// TIA Portal project "SSA-3GHz_V18" (V18) (continued)
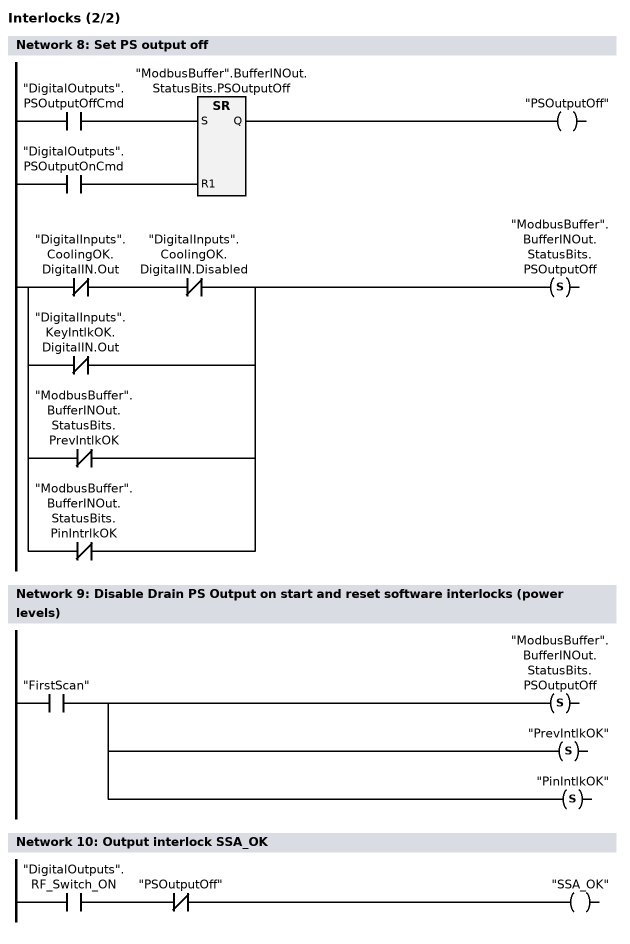
   RUNG wire#powerrail
      Contact( "DigitalOutputs".PSOutputOffCmd )
      S_SR(operand := "ModbusBuffer".BufferINOut.StatusBits.PSOutputOff, r1 := wire#w1)
      Coil( "PSOutputOff" )
   END_RUNG
   RUNG wire#powerrail
      Contact( "DigitalOutputs".PSOutputOnCmd )
   END_RUNG wire#w1
   RUNG wire#powerrail
      I_Contact( "DigitalInputs".CoolingOK.DigitalIN.Out )
      I_Contact( "DigitalInputs".CoolingOK.DigitalIN.Disabled )
      wire#w2
      S_Coil( "ModbusBuffer".BufferINOut.StatusBits.PSOutputOff )
   END_RUNG
   RUNG wire#powerrail
      I_Contact( "DigitalInputs".KeyIntlkOK.DigitalIN.Out )
   END_RUNG wire#w2
   RUNG wire#powerrail
      I_Contact( "ModbusBuffer".BufferINOut.StatusBits.PrevIntlkOK )
   END_RUNG wire#w2
   RUNG wire#powerrail
      I_Contact( "ModbusBuffer".BufferINOut.StatusBits.PinIntrlkOK )
   END_RUNG wire#w2
   // the same network as SCL:
   IF "DigitalOutputs".PSOutputOffCmd THEN
       "ModbusBuffer".BufferINOut.StatusBits.PSOutputOff := TRUE;   // SR flip-flop
   END_IF;
   IF "DigitalOutputs".PSOutputOnCmd THEN "ModbusBuffer".BufferINOut.StatusBits.PSOutputOff := FALSE; END_IF;
   "PSOutputOff" := "ModbusBuffer".BufferINOut.StatusBits.PSOutputOff;
   IF (NOT "DigitalInputs".CoolingOK.DigitalIN.Out AND NOT "DigitalInputs".CoolingOK.DigitalIN.Disabled) OR NOT "DigitalInputs".KeyIntlkOK.DigitalIN.Out OR NOT "ModbusBuffer".BufferINOut.StatusBits.PrevIntlkOK OR NOT "ModbusBuffer".BufferINOut.StatusBits.PinIntrlkOK THEN
       "ModbusBuffer".BufferINOut.StatusBits.PSOutputOff := TRUE;
   END_IF;
END_REGION

REGION Network 9: Disable Drain PS Output on start and reset software interlocks (power levels)
   RUNG wire#powerrail
      Contact( "FirstScan" )
      wire#w1
      S_Coil( "ModbusBuffer".BufferINOut.StatusBits.PSOutputOff )
   END_RUNG
   RUNG wire#w1
      S_Coil( "PrevIntlkOK" )
   END_RUNG
   RUNG wire#w1
      S_Coil( "PinIntlkOK" )
   END_RUNG
   // the same network as SCL:
   IF "FirstScan" THEN
       "ModbusBuffer".BufferINOut.StatusBits.PSOutputOff := TRUE;
       "PrevIntlkOK" := TRUE;
       "PinIntlkOK" := TRUE;
   END_IF;
END_REGION

REGION Network 10: Output interlock SSA_OK
   RUNG wire#powerrail
      Contact( "DigitalOutputs".RF_Switch_ON )
      I_Contact( "PSOutputOff" )
      Coil( "SSA_OK" )
   END_RUNG
   // the same network as SCL:
   "SSA_OK" := "DigitalOutputs".RF_Switch_ON AND NOT "PSOutputOff";
END_REGION
END_FUNCTION

ORGANIZATION_BLOCK "Main"   // OB1, LAD, ProgramCycle
TITLE = "Main Program Sweep (Cycle)"
{ S7_Optimized_Access := 'TRUE' }
VERSION : 0.1
   VAR_INPUT
      Initial_Call : Bool;   // Initial call of this OB
      Remanence : Bool;   // =True, if remanent data are available
   END_VAR
   VAR_TEMP
      trigger : Bool;   // 1 for one cycle
   END_VAR
BEGIN

REGION Network 1: Setup
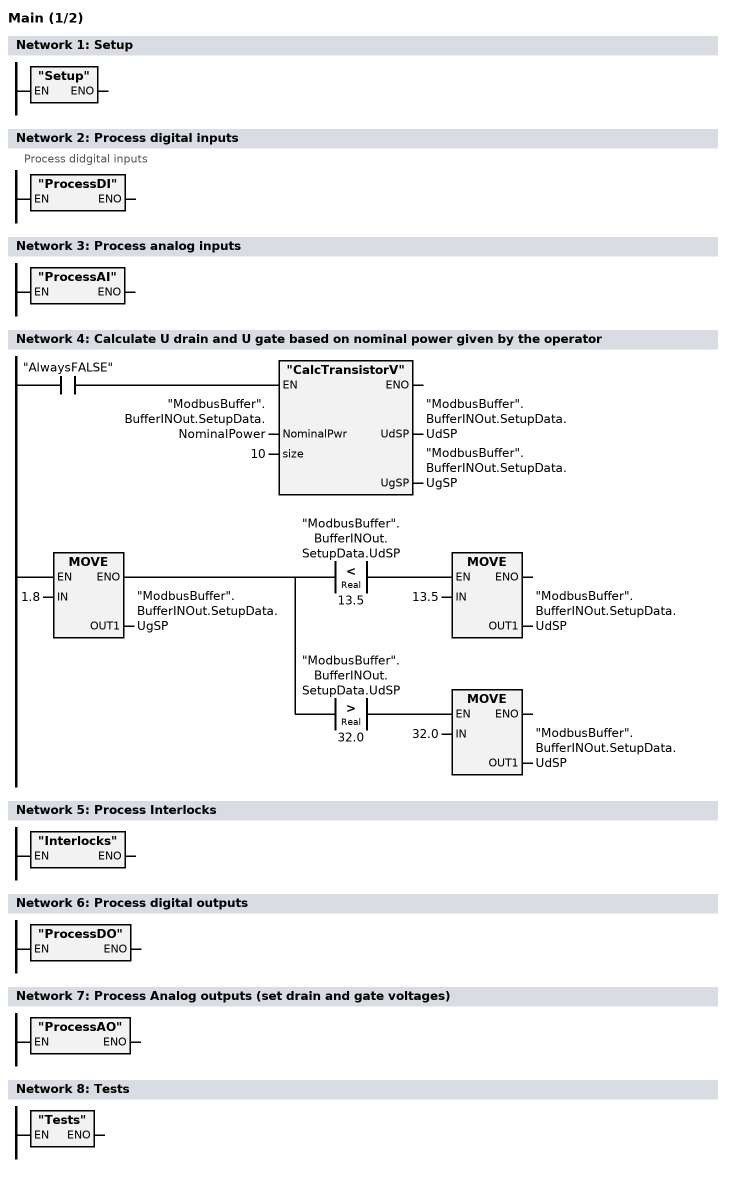
   RUNG wire#powerrail
      "Setup"()
   END_RUNG
   // the same network as SCL:
   "Setup"();
END_REGION

REGION Network 2: Process digital inputs
   // Process didgital inputs
   RUNG wire#powerrail
      "ProcessDI"()
   END_RUNG
   // the same network as SCL:
   "ProcessDI"();
END_REGION

REGION Network 3: Process analog inputs
   RUNG wire#powerrail
      "ProcessAI"()
   END_RUNG
   // the same network as SCL:
   "ProcessAI"();
END_REGION

REGION Network 4: Calculate U drain and U gate based on nominal power given by the operator
   RUNG wire#powerrail
      Contact( "AlwaysFALSE" )
      "CalcTransistorV"(NominalPwr := "ModbusBuffer".BufferINOut.SetupData.NominalPower, size := 10, UdSP => "ModbusBuffer".BufferINOut.SetupData.UdSP, UgSP => "ModbusBuffer".BufferINOut.SetupData.UgSP)
   END_RUNG
   RUNG wire#powerrail
      Move(in := 1.8, out1 => "ModbusBuffer".BufferINOut.SetupData.UgSP)
      wire#w1
      { S7_Templates := "SrcType := Real" } LT_Contact(in1 := "ModbusBuffer".BufferINOut.SetupData.UdSP, in2 := 13.5)
      Move(in := 13.5, out1 => "ModbusBuffer".BufferINOut.SetupData.UdSP)
   END_RUNG
   RUNG wire#w1
      { S7_Templates := "SrcType := Real" } GT_Contact(in1 := "ModbusBuffer".BufferINOut.SetupData.UdSP, in2 := 32.0)
      Move(in := 32.0, out1 => "ModbusBuffer".BufferINOut.SetupData.UdSP)
   END_RUNG
   // the same network as SCL:
   IF "AlwaysFALSE" THEN
       "CalcTransistorV"(NominalPwr := "ModbusBuffer".BufferINOut.SetupData.NominalPower,
                         size := 10,
                         UdSP => "ModbusBuffer".BufferINOut.SetupData.UdSP,
                         UgSP => "ModbusBuffer".BufferINOut.SetupData.UgSP);
   END_IF;
   "ModbusBuffer".BufferINOut.SetupData.UgSP := 1.8;
   IF "ModbusBuffer".BufferINOut.SetupData.UdSP < 13.5 THEN
       "ModbusBuffer".BufferINOut.SetupData.UdSP := 13.5;
   END_IF;
   IF "ModbusBuffer".BufferINOut.SetupData.UdSP > 32.0 THEN
       "ModbusBuffer".BufferINOut.SetupData.UdSP := 32.0;
   END_IF;
END_REGION

REGION Network 5: Process Interlocks
   RUNG wire#powerrail
      "Interlocks"()
   END_RUNG
   // the same network as SCL:
   "Interlocks"();
END_REGION

REGION Network 6: Process digital outputs
   RUNG wire#powerrail
      "ProcessDO"()
   END_RUNG
   // the same network as SCL:
   "ProcessDO"();
END_REGION

REGION Network 7: Process Analog outputs (set drain and gate voltages)
   RUNG wire#powerrail
      "ProcessAO"()
   END_RUNG
   // the same network as SCL:
   "ProcessAO"();
END_REGION

REGION Network 8: Tests
   RUNG wire#powerrail
      "Tests"()
   END_RUNG
   // the same network as SCL:
   "Tests"();
END_REGION

REGION Network 9: ModBus server
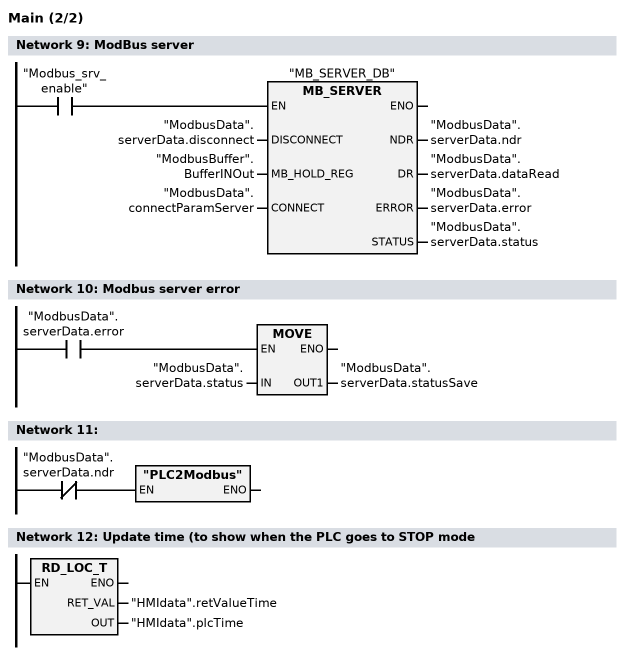
   IF "Modbus_srv_enable" THEN
       "MB_SERVER_DB"(DISCONNECT := "ModbusData".serverData.disconnect,   // MB_SERVER
                      MB_HOLD_REG := "ModbusBuffer".BufferINOut,
                      CONNECT := "ModbusData".connectParamServer,
                      NDR => "ModbusData".serverData.ndr,
                      DR => "ModbusData".serverData.dataRead,
                      ERROR => "ModbusData".serverData.error,
                      STATUS => "ModbusData".serverData.status);
   END_IF;
END_REGION

REGION Network 10: Modbus server error
   RUNG wire#powerrail
      Contact( "ModbusData".serverData.error )
      Move(in := "ModbusData".serverData.status, out1 => "ModbusData".serverData.statusSave)
   END_RUNG
   // the same network as SCL:
   IF "ModbusData".serverData.error THEN
       "ModbusData".serverData.statusSave := "ModbusData".serverData.status;
   END_IF;
END_REGION

REGION Network 11
   RUNG wire#powerrail
      I_Contact( "ModbusData".serverData.ndr )
      "PLC2Modbus"()
   END_RUNG
   // the same network as SCL:
   IF NOT "ModbusData".serverData.ndr THEN "PLC2Modbus"(); END_IF;
END_REGION

REGION Network 12: Update time (to show when the PLC goes to STOP mode
   "HMIdata".retValueTime := RD_LOC_T(OUT => "HMIdata".plcTime);
END_REGION
END_ORGANIZATION_BLOCK

// folder: 5_T_CONFIG (S7-1200, S7-1500)

FUNCTION_BLOCK "SLI_FB_T_CONFIG"   // FB4, LAD
{ S7_Optimized_Access := 'TRUE' }
VERSION : 0.1
// Info: The example is meant to change the PROFINET  device name and IP address of the CPU via its PROFINET interface.
   VAR
      T_CONFIG_Instance : T_CONFIG;
      done : Bool;
      errorLocation : DWord;
   END_VAR
BEGIN

REGION Network 1: Set "start" to TRUE to configure the PROFINET interface.
   // NOTE! Before using the example:
   // 
   // Condition:
   // 1) Open the device view of the CPU "> Properties > PROFINET interface > Ethernet addresses > PROFINET". 
   // 2) To set the device name: Activate the following options: 
   // - "IP address is set directly at the device". 
   // - "PROFINET device name is set directly at the device".
   // 
   // Regarding parameter INTERFACE ("hwid"):
   // - Change the value of "hwid" according to the identification number of the PROFINET interface of your local device (CPU). (Open "PLC tags > Show all tags > System constants. Look for a name like "<Local~PROFINET_interface_1>" with a Data type "Hw_Interface". The cell "value" contains the hwid.)
   // 
   // Info:
   // In the "header" (IF_CONF_HEADER):
   // - SubfieldCount = 2: Indicates that two additional structures ("deviceIP" and "deviceName") are used below.
   // 
   // In the structure "deviceIP" (system data type IF_CONF_v4):
   // - Lenght = 18: Information on overall length of the structure (12 bytes for the device IP + 6 bytes for the parameters Id, Length and Mode)
   // - Mode = 1: Permanent change of the device IP.
   // - InterfaceAddress, SubnetMask, DefaultRouter: IP connection data.
   // 
   // In the structure "deviceName" (system data type IF_CONF_NOS):
   // - Lenght = 11: Information on overall length of the structure (5 bytes for the device name "myplc" + 6 bytes for the parameters Id, Length and Mode)
   // - Mode = 1: Permanent change of the device name in "myplc".
   // - NOS[1] ... NOS[5]: Device name (1 character / byte)
   // 
   // Note: Instead of an absolute length, you can use the default start value (Lenght = 0) for a dynamic length.
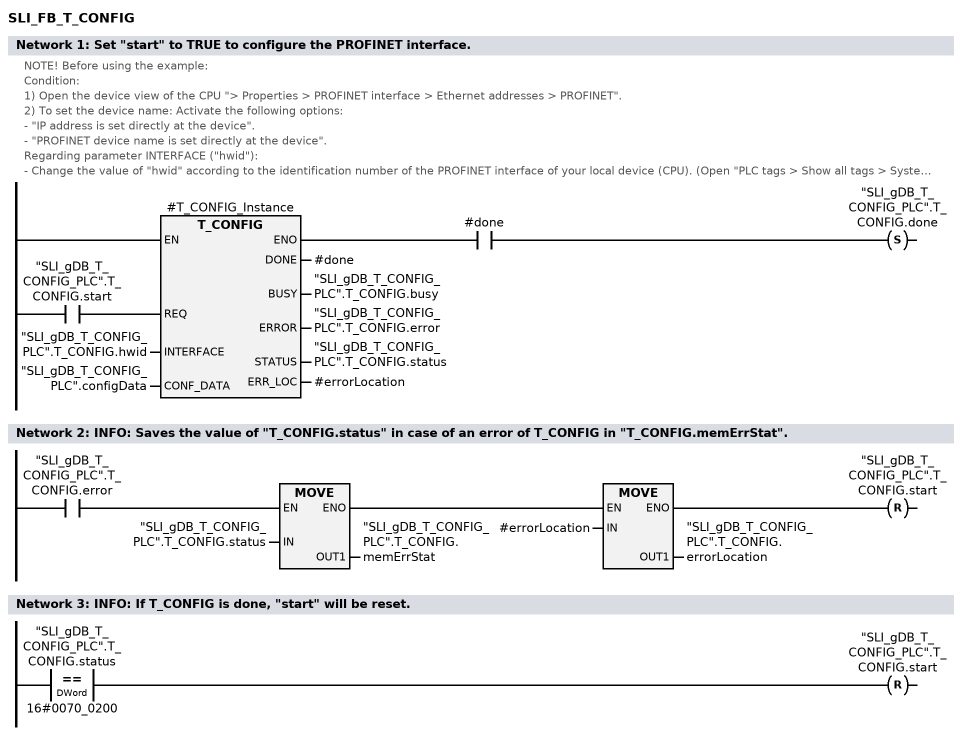
   // ENO of a box is taken as its EN; it also drops when the box reports an error
   #T_CONFIG_Instance(Req := "SLI_gDB_T_CONFIG_PLC".T_CONFIG.start,   // T_CONFIG
                      Interface := "SLI_gDB_T_CONFIG_PLC".T_CONFIG.hwid,
                      Conf_Data := "SLI_gDB_T_CONFIG_PLC".configData,
                      Done => #done,
                      Busy => "SLI_gDB_T_CONFIG_PLC".T_CONFIG.busy,
                      Error => "SLI_gDB_T_CONFIG_PLC".T_CONFIG.error,
                      Status => "SLI_gDB_T_CONFIG_PLC".T_CONFIG.status,
                      Err_Loc => #errorLocation);
   IF #done THEN "SLI_gDB_T_CONFIG_PLC".T_CONFIG.done := TRUE; END_IF;
END_REGION

REGION Network 2: INFO: Saves the value of "T_CONFIG.status" in case of an error of T_CONFIG in "T_CONFIG.memErrStat".
   RUNG wire#powerrail
      Contact( "SLI_gDB_T_CONFIG_PLC".T_CONFIG.error )
      Move(in := "SLI_gDB_T_CONFIG_PLC".T_CONFIG.status, out1 => "SLI_gDB_T_CONFIG_PLC".T_CONFIG.memErrStat)
      Move(in := #errorLocation, out1 => "SLI_gDB_T_CONFIG_PLC".T_CONFIG.errorLocation)
      R_Coil( "SLI_gDB_T_CONFIG_PLC".T_CONFIG.start )
   END_RUNG
   // the same network as SCL:
   IF "SLI_gDB_T_CONFIG_PLC".T_CONFIG.error THEN
       "SLI_gDB_T_CONFIG_PLC".T_CONFIG.memErrStat := "SLI_gDB_T_CONFIG_PLC".T_CONFIG.status;
       "SLI_gDB_T_CONFIG_PLC".T_CONFIG.errorLocation := #errorLocation;
       "SLI_gDB_T_CONFIG_PLC".T_CONFIG.start := FALSE;
   END_IF;
END_REGION

REGION Network 3: INFO: If T_CONFIG is done, "start" will be reset.
   RUNG wire#powerrail
      { S7_Templates := "SrcType := DWord" } EQ_Contact(in1 := "SLI_gDB_T_CONFIG_PLC".T_CONFIG.status, in2 := 16#0070_0200)
      R_Coil( "SLI_gDB_T_CONFIG_PLC".T_CONFIG.start )
   END_RUNG
   // the same network as SCL:
   IF "SLI_gDB_T_CONFIG_PLC".T_CONFIG.status = 16#0070_0200 THEN
       "SLI_gDB_T_CONFIG_PLC".T_CONFIG.start := FALSE;
   END_IF;
END_REGION
END_FUNCTION_BLOCK

(* ===== HMI "HMI_RT_1" =====
system functions are stored by id; their names below are inferred from use
connection "HMI_Connection_1": ETHERNET, SMART_S7_1200_OMS

HMI tags "Default tag table"
   "Tag_ScreenNumber" : UInt, internal
   "AnalogInputs_Pfwd_AnalogIN_Out" : Real = PLC AnalogInputs.Pfwd.AnalogIN.Out, 1 s
   "AnalogInputs_Prev_AnalogIN_Out" : Real = PLC AnalogInputs.Prev.AnalogIN.Out, 1 s
   "DigitalInputs_DutyCycOK_DigitalIN_Out" : Bool = PLC DigitalInputs.DutyCycOK.DigitalIN.Out, 1 s
   "DigitalInputs_KeyIntlkOK_DigitalIN_Out" : Bool = PLC DigitalInputs.KeyIntlkOK.DigitalIN.Out, 1 s
   "DigitalInputs_ExtIntlkT1_DigitalIN_Out" : Bool = PLC DigitalInputs.ExtIntlk1.DigitalIN.Out, 1 s
   "DigitalInputs_ExtIntlkT3_DigitalIN_Out" : Bool = PLC DigitalInputs.ExtIntlk2.DigitalIN.Out, 1 s
   "AnalogInputs_U_drain_RBK_AnalogIN_Out" : Real = PLC AnalogInputs.U_drain_RBK.AnalogIN.Out, 1 s
   "AnalogInputs_Pin_AnalogIN_Out" : Real = PLC AnalogInputs.Pin.AnalogIN.Out, 1 s
   "StatusBits_T1_OK_DigitalIN_Out" : Bool = PLC ModbusBuffer.BufferINOut.StatusBits.T1_OK AT %DB101.DBX208.4, 1 s
   "DigitalInputs_CoolingWtrOK_DigitalIN_Out" : Bool = PLC DigitalInputs.CoolingOK.DigitalIN.Out, 1 s
   "DigitalInputs_SoftIntlk1_DigitalIN_Out" : Bool = PLC DigitalInputs.SofIntlk1.DigitalIN.Out, 1 s
   "DigitalInputs_SoftIntlk2_DigitalIN_Out" : Bool = PLC DigitalInputs.SoftIntlk2.DigitalIN.Out, 1 s
   "TestBlink" : Bool = PLC TestBlink AT %Q1.0, 1 s
   "AnalogInputs_U_gate_RBK_AnalogIN_VisuState" : Byte = PLC AnalogInputs.Pin.AnalogIN.VisuState, 1 s
   "VisuTest" : Byte = PLC VisuTest AT %MB104, 1 s
   "DigitalInputs_DutyCycOK_DigitalIN_Disabled" : Bool = PLC DigitalInputs.DutyCycOK.DigitalIN.Disabled, 1 s
   "DigitalInputs_KeyIntlkOK_DigitalIN_Disabled" : Bool = PLC DigitalInputs.KeyIntlkOK.DigitalIN.Disabled, 1 s
   "DigitalInputs_ExtIntlk1_DigitalIN_Disabled" : Bool = PLC DigitalInputs.ExtIntlk1.DigitalIN.Disabled, 1 s
   "DigitalInputs_ExtIntlk2_DigitalIN_Disabled" : Bool = PLC DigitalInputs.ExtIntlk2.DigitalIN.Disabled, 1 s
   "DigitalInputs_T1_OK_DigitalIN_Disabled" : Bool = PLC DigitalInputs.T1_OK.DigitalIN.Disabled, 1 s
   "DigitalInputs_CoolingOK_DigitalIN_Disabled" : Bool = PLC DigitalInputs.CoolingOK.DigitalIN.Disabled, 1 s
   "DigitalInputs_SoftIntlk1_DigitalIN_Disabled" : Bool = PLC DigitalInputs.SofIntlk1.DigitalIN.Disabled, 1 s
   "DigitalInputs_SoftIntlk2_DigitalIN_Disabled" : Bool = PLC DigitalInputs.SoftIntlk2.DigitalIN.Disabled, 1 s
   "ModbusBuffer_BufferINOut_SetupData_RemoteMode" : Bool = PLC ModbusBuffer.BufferINOut.SetupData.RemoteMode AT %DB101.DBX120.0, 1 s
   "ModbusBuffer_BufferINOut_SetupData_NominalPower" : Real = PLC ModbusBuffer.BufferINOut.SetupData.NominalPower AT %DB101.DBD122, 1 s
   "Counter_HMI" : UDInt = PLC Counter AT %MD100, 1 s
   "SLI_gDB_T_CONFIG_PLC_configData_deviceIP_InterfaceAddress_ADDR{1}" : Byte = PLC SLI_gDB_T_CONFIG_PLC.configData.deviceIP.InterfaceAddress.ADDR[1], 1 s
   "SLI_gDB_T_CONFIG_PLC_configData_deviceIP_InterfaceAddress_ADDR{2}" : Byte = PLC SLI_gDB_T_CONFIG_PLC.configData.deviceIP.InterfaceAddress.ADDR[2], 1 s
   "SLI_gDB_T_CONFIG_PLC_configData_deviceIP_InterfaceAddress_ADDR{3}" : Byte = PLC SLI_gDB_T_CONFIG_PLC.configData.deviceIP.InterfaceAddress.ADDR[3], 1 s
   "SLI_gDB_T_CONFIG_PLC_configData_deviceIP_InterfaceAddress_ADDR{4}" : Byte = PLC SLI_gDB_T_CONFIG_PLC.configData.deviceIP.InterfaceAddress.ADDR[4], 1 s
   "IP_SubnetMask_ADDR{1}" : Byte = PLC SLI_gDB_T_CONFIG_PLC.configData.deviceIP.SubnetMask.ADDR[1] AT %DB1.DBB0, 1 s
   "IP_SubnetMask_ADDR{2}" : Byte = PLC SLI_gDB_T_CONFIG_PLC.configData.deviceIP.SubnetMask.ADDR[2] AT %DB1.DBB0, 1 s
   "IP_SubnetMask_ADDR{3}" : Byte = PLC SLI_gDB_T_CONFIG_PLC.configData.deviceIP.SubnetMask.ADDR[3] AT %DB1.DBB0, 1 s
   "IP_SubnetMask_ADDR{4}" : Byte = PLC SLI_gDB_T_CONFIG_PLC.configData.deviceIP.SubnetMask.ADDR[4] AT %DB1.DBB0, 1 s
   "IP_DefaultRouter_ADDR{1}" : Byte = PLC SLI_gDB_T_CONFIG_PLC.configData.deviceIP.DefaultRouter.ADDR[1] AT %DB1.DBB0, 1 s
   "IP_DefaultRouter_ADDR{2}" : Byte = PLC SLI_gDB_T_CONFIG_PLC.configData.deviceIP.DefaultRouter.ADDR[2] AT %DB1.DBB0, 1 s
   "IP_DefaultRouter_ADDR{3}" : Byte = PLC SLI_gDB_T_CONFIG_PLC.configData.deviceIP.DefaultRouter.ADDR[3] AT %DB1.DBB0, 1 s
   "IP_DefaultRouter_ADDR{4}" : Byte = PLC SLI_gDB_T_CONFIG_PLC.configData.deviceIP.DefaultRouter.ADDR[4] AT %DB1.DBB0, 1 s
   "Set_IP_PArameters" : Bool = PLC Set_IP_PArameters AT %M10.2, 1 s
   "evaluationLiveBit" : Bool AT %DB103.DBX1.2, 1 s
      on ChangeValue: function_c655a98f("HMI_Connection_1", "HMIdata_getPlcMode")
   "hmi_plcTime" : DTL = PLC HMIdata.plcTime AT %DB103.DBX4.0, 1 s
   "HMIdata_getPlcMode" : Int = PLC HMIdata.getPlcMode AT %DB103.DBW2, 1 s
   "ModbusBuffer_BufferINOut_SetupData_dBm_unit" : Bool = PLC ModbusBuffer.BufferINOut.SetupData.dBm_unit AT %DB101.DBX120.1, 1 s
   "ModbusBuffer_BufferINOut_CalculatedData_Pfwd_dBm" : Real = PLC ModbusBuffer.BufferINOut.CalculatedData.Pfwd_dBm AT %DB101.DBD180, 1 s
   "ModbusBuffer_BufferINOut_CalculatedData_Prev_dBm" : Real = PLC ModbusBuffer.BufferINOut.CalculatedData.Prev_dBm AT %DB101.DBD184, 1 s
   "ModbusBuffer_BufferINOut_SetupData_NominalPower_dBm" : Real = PLC ModbusBuffer.BufferINOut.SetupData.NominalPower_dBm AT %DB101.DBD126, 1 s
   "ModbusBuffer_BufferINOut_ADCdata_TT01" : Real = PLC ModbusBuffer.BufferINOut.ADCdata.TT01 AT %DB101.DBD164, 1 s
   "ModbusBuffer_BufferINOut_ADCdata_TT04" : Real = PLC ModbusBuffer.BufferINOut.ADCdata.TT04 AT %DB101.DBD176, 1 s
   "ModbusBuffer_BufferINOut_ADCdata_TT03" : Real = PLC ModbusBuffer.BufferINOut.ADCdata.TT03 AT %DB101.DBD172, 1 s
   "ModbusBuffer_BufferINOut_ADCdata_TT02" : Real = PLC ModbusBuffer.BufferINOut.ADCdata.TT02 AT %DB101.DBD168, 1 s
   "ModbusBuffer_BufferINOut_Commands_Reset" : Bool = PLC ModbusBuffer.BufferINOut.Commands.Reset AT %DB101.DBX138.3, 1 s
   "HMI_Tag_Efficiency" : Real = PLC ModbusBuffer.BufferINOut.CalculatedData.Effic AT %DB101.DBD188, 1 s
   "RFSwitchStatus" : Bool = PLC ModbusBuffer.BufferINOut.StatusBits.RFSwitchON AT %DB101.DBX210.0, 1 s
   "ModbusBuffer_BufferINOut_CalculatedData_AmplVisuState" : Byte = PLC ModbusBuffer.BufferINOut.CalculatedData.AmplVisuState AT %DB101.DBB196, 1 s
   "ModbusBuffer_BufferINOut_Commands_PSOutputOn" : Bool = PLC ModbusBuffer.BufferINOut.Commands.PSOutputOn AT %DB101.DBX138.0, 1 s
   "ModbusBuffer_BufferINOut_Commands_PSOutputOff" : Bool = PLC ModbusBuffer.BufferINOut.Commands.PSOutputOff AT %DB101.DBX138.1, 1 s
   "ModbusBuffer_BufferINOut_CalculatedData_Prev_dBm(1)" : Real = PLC ModbusBuffer.BufferINOut.CalculatedData.Prev_dBm AT %DB101.DBD184, 1 s
   "ModbusBuffer_BufferINOut_SetupData_UdSP" : Real = PLC ModbusBuffer.BufferINOut.SetupData.UdSP AT %DB101.DBD130, 1 s
   "RestoreFactorySettings" : Bool = PLC RestoreFactorySettings AT %M10.7, 1 s
   "ModbusBuffer_BufferINOut_CalculatedData_Pin_dBm" : Real = PLC ModbusBuffer.BufferINOut.CalculatedData.Pin_dBm AT %DB101.DBD192, 1 s
   "ModbusBuffer_BufferINOut_LookupTable_PinA" : Real = PLC ModbusBuffer.BufferINOut.LookupTable.PinA AT %DB101.DBD96, 1 s
   "ModbusBuffer_BufferINOut_LookupTable_PinB" : Real = PLC ModbusBuffer.BufferINOut.LookupTable.PinB AT %DB101.DBD100, 1 s
   "ModbusBuffer_BufferINOut_LookupTable_PfwdA" : Real = PLC ModbusBuffer.BufferINOut.LookupTable.PfwdA AT %DB101.DBD112, 1 s
   "ModbusBuffer_BufferINOut_LookupTable_PfwdB" : Real = PLC ModbusBuffer.BufferINOut.LookupTable.PfwdB AT %DB101.DBD116, 1 s
   "ModbusBuffer_BufferINOut_LookupTable_PrevA" : Real = PLC ModbusBuffer.BufferINOut.LookupTable.PrevA AT %DB101.DBD104, 1 s
   "ModbusBuffer_BufferINOut_LookupTable_PrevB" : Real = PLC ModbusBuffer.BufferINOut.LookupTable.PrevB AT %DB101.DBD108, 1 s
   "ModbusBuffer_BufferINOut_PinLimitdBm" : Real = PLC ModbusBuffer.BufferINOut.PinLimitdBm AT %DB101.DBD216, 1 s
   "ModbusBuffer_BufferINOut_PrevFactor" : Real = PLC ModbusBuffer.BufferINOut.PrevFactor AT %DB101.DBD212, 1 s
   "PinUR" : Bool = PLC PinUR AT %M11.0, 1 s
   "PfwdUR" : Bool = PLC PfwdUR AT %M11.1, 1 s
   "PrevUR" : Bool = PLC PrevUR AT %M11.2, 1 s
   "ModbusBuffer_BufferINOut_StatusBits_SSA_OK" : Bool = PLC ModbusBuffer.BufferINOut.StatusBits.SSA_OK AT %DB101.DBX210.2, 1 s

text list "Text_list_loc_rem": 0 'To Rem.'; 1 'To Loc.'

text list "Text_list_EGU": 0 'W'; 1 'dBm'

text list "Textlist_GetPLCMode": 4 'SPS in STOP / STOP'; 8 'SPS in RUN / RUN'

text list "Text_list_underrange": 0 ''; 1 '<'

graphic list "Amplifier": 0 'Amplifier_grey_3'; 1 'Amplifier_blue_2'; 2 'Amplifier_green_2'; 3 'Amplifier_yellow_4'; 4 'Amplifier_red_3'

Template "Template" 480x272
   TextField "Template_Text field_1" at 94,6 size 23x37; Text 'P'
   TextField "Template_Text field_3" at 109,23 size 30x17; Text 'FWD'
   TextField "Template_Text field_5" at 291,8 size 23x37; Text 'P'
   TextField "Template_Text field_4" at 310,23 size 26x17; Text 'REV'
   Button "Alarms" at 1,46 size 63x44; TextOff 'Alarms'; PictureOff "AlarmDisplay_KTP400_Basic_PN_TR"; PictureOn "AlarmDisplay_KTP400_Basic_PN_TR"
      on Release: function_ef3f5d25("Alarm window_Unacknowledged", -1)
   Button "Start screen" at 1,226 size 63x44; TextOff 'Start screen'; PictureOff "NavigateHome_KTP400_Basic_PN_TR"; PictureOn "NavigateHome_KTP400_Basic_PN_TR"
      on Release: ActivateScreen("Root screen", 0)
   GraphicView "Logo" at 0,0 size 94x45; Picture "Logo of HMI_1"
   Button "Template_Button_3" at 1,91 size 63x44; TextOff 'System'
      on Release: ActivateScreen("System screens", 0)
   Group "Group" at 94,6 size 45x37
   Group "Group_1" at 291,8 size 45x37
   IOField "Template_I/O Pfwd" at 142,6 size 80x39; FormatPattern 999
      ProcessValue <- "AnalogInputs_Pfwd_AnalogIN_Out"
      Visibility <- "ModbusBuffer_BufferINOut_SetupData_dBm_unit"
   IOField "Template_I/O Prev" at 339,6 size 80x39; FormatPattern 999
      ProcessValue <- "AnalogInputs_Prev_AnalogIN_Out"
      Visibility <- "ModbusBuffer_BufferINOut_SetupData_dBm_unit"
   Switch "Template_Switch_1" at 1,136 size 64x44; CaptionText 'Switch'; TextOff 'Loc'; TextOn 'Rem'
      ProcessValue <- "ModbusBuffer_BufferINOut_SetupData_RemoteMode"
   Switch "Template_Switch_2" at 1,181 size 63x44; CaptionText 'Switch'; TextOff 'W'; TextOn 'dBm'
      ProcessValue <- "ModbusBuffer_BufferINOut_SetupData_dBm_unit"
   SymbolicIOField "Template_Symbolic I/O field_1" at 225,15 size 50x28; TextOff '0'; TextOn '1'; TextList "Text_list_EGU"
      ProcessValue <- "ModbusBuffer_BufferINOut_SetupData_dBm_unit"
   SymbolicIOField "Template_Symbolic I/O field_2" at 422,15 size 50x28; TextOn '1'; TextOff '0'; TextList "Text_list_EGU"
      ProcessValue <- "ModbusBuffer_BufferINOut_SetupData_dBm_unit"
   IOField "Template_I/O Pfwd dBm" at 142,6 size 80x39; FormatPattern 999.9
      Visibility <- "ModbusBuffer_BufferINOut_SetupData_dBm_unit"
      ProcessValue <- "ModbusBuffer_BufferINOut_CalculatedData_Pfwd_dBm"
   IOField "Template_I/O Prev dBm" at 339,6 size 80x39; FormatPattern 999.9
      Visibility <- "ModbusBuffer_BufferINOut_SetupData_dBm_unit"
      ProcessValue <- "ModbusBuffer_BufferINOut_CalculatedData_Prev_dBm"
   SymbolicIOField "Symbolic I/O Underrange Pfwd" at 140,5 size 22x39; TextOn '1'; TextOff '0'; TextList "Text_list_underrange"
      ProcessValue <- "PfwdUR"
   SymbolicIOField "Symbolic I/O Underrange Prev" at 337,5 size 22x39; TextOn '1'; TextOff '0'; TextList "Text_list_underrange"
      ProcessValue <- "PrevUR"

screen "Root screen" 480x272, template "Template_noPrev"
   on GenerateScreen: SetTag("Tag_ScreenNumber", 1)
   TextField "Text field_1" at 69,206 size 87x20; Text 'Interlocks In'
   TextField "Text field_2" at 74,227 size 75x20; Text 'Duty Cyc.'
      Appearance <- "DigitalInputs_DutyCycOK_DigitalIN_Out"
      Visibility <- "DigitalInputs_DutyCycOK_DigitalIN_Disabled"
   TextField "Text field_3" at 74,248 size 75x20; Text 'KeyIntlk'
      Appearance <- "DigitalInputs_KeyIntlkOK_DigitalIN_Out"
      Visibility <- "DigitalInputs_KeyIntlkOK_DigitalIN_Disabled"
   TextField "Text field_4" at 151,227 size 75x20; Text 'Ext Intlk1'
      Appearance <- "DigitalInputs_ExtIntlkT1_DigitalIN_Out"
      Visibility <- "DigitalInputs_ExtIntlk1_DigitalIN_Disabled"
   TextField "Text field_5" at 151,248 size 75x20; Text 'ExtIntlk2'
      Appearance <- "DigitalInputs_ExtIntlkT3_DigitalIN_Out"
      Visibility <- "DigitalInputs_ExtIntlk2_DigitalIN_Disabled"
   Group "Group" at 71,82 size 19x20
   Group "Group_1" at 64,166 size 25x25
   TextField "Text field_13" at 228,227 size 75x20; Text 'T1_OK'
      Appearance <- "StatusBits_T1_OK_DigitalIN_Out"
      Visibility <- "DigitalInputs_T1_OK_DigitalIN_Disabled"
   TextField "Text field_14" at 228,248 size 75x20; Text 'Cooling'
      Visibility <- "DigitalInputs_CoolingOK_DigitalIN_Disabled"
      Appearance <- "DigitalInputs_CoolingWtrOK_DigitalIN_Out"
   TextField "Text field_15" at 305,227 size 75x20; Text 'P rev'
      Appearance <- "DigitalInputs_SoftIntlk1_DigitalIN_Out"
      Visibility <- "DigitalInputs_SoftIntlk1_DigitalIN_Disabled"
   TextField "Text field_16" at 305,248 size 75x20; Text 'P in'
      Appearance <- "DigitalInputs_SoftIntlk2_DigitalIN_Out"
      Visibility <- "DigitalInputs_SoftIntlk2_DigitalIN_Disabled"
   TextField "Text field_17" at 75,131 size 37x20; Text 'RF In'
   TextField "Text field_18" at 408,133 size 47x20; Text 'RF Out'
   GraphicIOField "Graphic I/O field_2" at 181,79 size 175x128; PictureList "Amplifier"
      ProcessValue <- "ModbusBuffer_BufferINOut_CalculatedData_AmplVisuState"
   Group "Group_TT01" at 365,53 size 102x21; FormatPattern 9.9
   Group "Group_TT01_2" at 365,72 size 102x21; FormatPattern 9.9
   SymbolicIOField "Template_Symbolic I/O field_1" at 138,164 size 50x28; TextOn '1'; TextOff '0'; TextList "Text_list_EGU"
      ProcessValue <- "ModbusBuffer_BufferINOut_SetupData_dBm_unit"
   IOField "Template_I/O Pin W" at 89,168 size 50x20; FormatPattern 9.999
      Visibility <- "ModbusBuffer_BufferINOut_SetupData_dBm_unit"
      ProcessValue <- "AnalogInputs_Pin_AnalogIN_Out"
   IOField "U drain ADC" at 136,83 size 41x18; FormatPattern 99.9
      ProcessValue <- "AnalogInputs_U_drain_RBK_AnalogIN_Out"
   TextField "Text field_26" at 87,62 size 84x17; Text 'SetPoint RBK'
   TextField "Text field_33" at 392,227 size 75x20; Text 'SSA_OK'
      Appearance <- "ModbusBuffer_BufferINOut_StatusBits_SSA_OK"
   TextField "Text field_27" at 382,204 size 90x20; Text 'Interlock Out'
   TextField "Text field_8" at 71,82 size 14x20; Text 'V'
   TextField "Text field_10" at 79,88 size 11x14; Text 'D'
   TextField "Text field_9" at 64,166 size 16x25; Text 'P'
   TextField "Text field_12" at 74,176 size 15x14; Text 'IN'
   GraphicIOField "Graphic I/O field_1" at 125,131 size 45x23; PictureOff "JS Disconnecting Switch Off-RED"; PictureOn "JS Disconnecting Switch On-GREEN"
      ProcessValue <- "RFSwitchStatus"
   IOField "I/O U drain" at 95,78 size 44x28; FormatPattern 99.9
      ProcessValue <- "ModbusBuffer_BufferINOut_SetupData_UdSP"
   IOField "Template_I/O Pin dBm" at 89,168 size 50x20; FormatPattern 999.9
      Visibility <- "ModbusBuffer_BufferINOut_SetupData_dBm_unit"
      ProcessValue <- "ModbusBuffer_BufferINOut_CalculatedData_Pin_dBm"
   TextField "Text field_7" at 365,53 size 40x20; Text 'TT01:'
   IOField "I/O field_1" at 397,53 size 53x21; FormatPattern s99.9
      ProcessValue <- "ModbusBuffer_BufferINOut_ADCdata_TT01"
   TextField "Text field_19" at 447,53 size 20x20; Text '°C'
   TextField "Text field_22" at 365,72 size 40x20; Text 'TT02:'
   IOField "I/O field_6" at 397,72 size 53x21; FormatPattern 99.9
      ProcessValue <- "ModbusBuffer_BufferINOut_ADCdata_TT02"
   TextField "Text field_23" at 447,72 size 20x20; Text '°C'
   SymbolicIOField "Template_Symbolic I/O Underrange" at 89,168 size 22x20; TextOn '1'; TextOff '0'; TextList "Text_list_underrange"
      ProcessValue <- "PinUR"

screen "System screens" 480x272, template "Template"
   on GenerateScreen: SetTag("Tag_ScreenNumber", 2)
   TextField "HmiScreenItemData" at 223,46 size 123x22; Text 'System screens'
   Button "Back" at 65,46 size 136x30; TextOff 'Back'
      on Release: ActivateScreen("Root screen", 0)
   Button "SIMATIC PLC system diagnostics" at 65,77 size 136x30; TextOff 'SIMATIC PLC s...'
      on Release: ActivateScreen("SIMATIC PLC system diagnostics", 0)
   Button "Project information" at 65,108 size 136x30; TextOff 'Calibrations...'; TextOn 'Project informat...'
      on Release: ActivateScreen("Calibrations", 0)
   Button "System information" at 65,139 size 136x30; TextOff 'System informa...'
      on Release: ActivateScreen("System information", 0)
   Button "Button_7" at 291,70 size 78x32; TextOn 'PLC STOP'; TextOff 'PLC STOP'
      on Release: function_f249594b("HMI_Connection_1", 4)
   Button "Button_6" at 208,70 size 79x32; TextOn 'PLC RUN'; TextOff 'PLC RUN'
      on Release: function_f249594b("HMI_Connection_1", 8)
   TextField "Text field_1" at 79,186 size 85x20; Text 'PLC IP Addr.'
   TextField "Text field_2" at 80,214 size 82x20; Text 'PLC IP Mask'
   TextField "Text field_3" at 88,238 size 62x20; Text 'Gateway'
   Group "Group_3" at 175,175 size 177x36
   Group "Group_7" at 175,206 size 177x36
   Group "Group_11" at 175,236 size 177x36
   Button "Button_1" at 359,224 size 115x43; TextOff 'Load the new network settings'
      on Release: SetBit("Set_IP_PArameters")
   Button "Button_2" at 358,175 size 116x44; TextOff 'Stop HMI RunTime'
      on Release: StopRuntime(0)
   IOField "I/O field_13" at 289,123 size 181x32; FormatPattern 9999999999999999999999999999999999999999
      ProcessValue <- "hmi_plcTime"
   Button "Button_3" at 373,70 size 96x49; TextOff 'Screen Calibration'
      on Click: function_bc3e350c()
   Button "Button_Restore_inactive" at 208,108 size 80x62; HelpText 'Active only in Local mode Restore Ud look-up table. IP addr. 192.168.1.234/24 Gateway: 192.168.1.1'; TextOff 'Restore Factory Settings'
   Button "Button_Restore_active" at 208,108 size 80x62; TextOff 'Restore Factory Settings'; HelpText 'Restore Ud look-up table. IP addr. 192.168.1.234/24 Gateway: 192.168.1.1'
      on Release: ResetBit("RestoreFactorySettings")
      on Press: SetBit("RestoreFactorySettings")
      Visibility <- "ModbusBuffer_BufferINOut_SetupData_RemoteMode"
   IOField "I/O field_1" at 175,175 size 39x32; FormatPattern 999
      ProcessValue <- "SLI_gDB_T_CONFIG_PLC_configData_deviceIP_InterfaceAddress_ADDR{1}"
   TextField "Text field_4" at 211,184 size 11x27; Text '.'
   Group "Group" at 175,175 size 47x36
   Group "Group_1" at 221,175 size 47x36
   Group "Group_2" at 267,175 size 47x36
   IOField "I/O field_4" at 313,175 size 39x32; FormatPattern 999
      ProcessValue <- "SLI_gDB_T_CONFIG_PLC_configData_deviceIP_InterfaceAddress_ADDR{4}"
   IOField "I/O field_2" at 221,175 size 39x32; FormatPattern 999
      ProcessValue <- "SLI_gDB_T_CONFIG_PLC_configData_deviceIP_InterfaceAddress_ADDR{2}"
   TextField "Text field_5" at 257,184 size 11x27; Text '.'
   IOField "I/O field_3" at 267,175 size 39x32; FormatPattern 999
      ProcessValue <- "SLI_gDB_T_CONFIG_PLC_configData_deviceIP_InterfaceAddress_ADDR{3}"
   TextField "Text field_6" at 303,184 size 11x27; Text '.'
   IOField "I/O field_5" at 175,206 size 39x32; FormatPattern 999
      ProcessValue <- "IP_SubnetMask_ADDR{1}"
   TextField "Text field_7" at 211,215 size 11x27; Text '.'
   Group "Group_4" at 175,206 size 47x36
   Group "Group_5" at 221,206 size 47x36
   Group "Group_6" at 267,206 size 47x36
   IOField "I/O field_8" at 313,206 size 39x32; FormatPattern 999
      ProcessValue <- "IP_SubnetMask_ADDR{4}"
   IOField "I/O field_6" at 221,206 size 39x32; FormatPattern 999
      ProcessValue <- "IP_SubnetMask_ADDR{2}"
   TextField "Text field_8" at 257,215 size 11x27; Text '.'
   IOField "I/O field_7" at 267,206 size 39x32; FormatPattern 999
      ProcessValue <- "IP_SubnetMask_ADDR{3}"
   TextField "Text field_9" at 303,215 size 11x27; Text '.'
   IOField "I/O field_9" at 175,236 size 39x32; FormatPattern 999
      ProcessValue <- "IP_DefaultRouter_ADDR{1}"
   TextField "Text field_10" at 211,245 size 11x27; Text '.'
   Group "Group_8" at 175,236 size 47x36
   Group "Group_9" at 221,236 size 47x36
   Group "Group_10" at 267,236 size 47x36
   IOField "I/O field_12" at 313,236 size 39x32; FormatPattern 999
      ProcessValue <- "IP_DefaultRouter_ADDR{4}"
   IOField "I/O field_10" at 221,236 size 39x32; FormatPattern 999
      ProcessValue <- "IP_DefaultRouter_ADDR{2}"
   TextField "Text field_11" at 257,245 size 11x27; Text '.'
   IOField "I/O field_11" at 267,236 size 39x32; FormatPattern 999
      ProcessValue <- "IP_DefaultRouter_ADDR{3}"
   TextField "Text field_12" at 303,245 size 11x27; Text '.'

screen "SIMATIC PLC system diagnostics" 480x272, template "Template"
   on GenerateScreen: SetTag("Tag_ScreenNumber", 3)
   SysDiagControl "HmiScreenItemData" at 65,77 size 412x188
   Button "Back" at 65,46 size 136x30; TextOff 'Back'
      on Release: ActivateScreen("System screens", 0)

screen "Calibrations" 480x272, template "Template"
   on GenerateScreen: SetTag("Tag_ScreenNumber", 4)
   TextField "Text field_1" at 78,56 size 228x68; Text 'Calibration constants A and B for the power measurements U is the voltage on the ADC input P[dBm]=A[dBm/V]*U[V]+B[dBm]'
   TextField "Text field_5" at 142,130 size 90x20; Text 'A B'
   Group "Pin" at 78,150 size 170x32
   Group "Pfwd" at 78,186 size 170x32
   Group "Prev" at 78,222 size 170x32
   TextField "Text field_6" at 328,56 size 132x20; Text 'Interlock constants'
   TextField "Text field_7" at 312,102 size 102x20; Text 'Pin Max [dBm]:'
   TextField "Text field_8" at 312,138 size 110x20; Text 'Prev/Pfwd Max:'
   IOField "I/O field_7" at 422,96 size 52x32; FormatPattern 99.9
      ProcessValue <- "ModbusBuffer_BufferINOut_PinLimitdBm"
   IOField "I/O field_8" at 422,132 size 52x32; FormatPattern 9.99
      ProcessValue <- "ModbusBuffer_BufferINOut_PrevFactor"
   Group "Group_1" at 340,224 size 32x25
   SymbolicIOField "Template_Symbolic I/O field_1" at 421,224 size 50x28; TextOn '1'; TextOff '0'; TextList "Text_list_EGU"
      ProcessValue <- "ModbusBuffer_BufferINOut_SetupData_dBm_unit"
   IOField "Template_I/O Pin W" at 372,228 size 50x20; FormatPattern 9.999
      Visibility <- "ModbusBuffer_BufferINOut_SetupData_dBm_unit"
      ProcessValue <- "AnalogInputs_Prev_AnalogIN_Out"
   TextField "Text field_2" at 78,156 size 45x20; Text 'Pin:'
   IOField "I/O field_1" at 122,150 size 59x32; FormatPattern 99.99
      ProcessValue <- "ModbusBuffer_BufferINOut_LookupTable_PinA"
   IOField "I/O field_2" at 185,150 size 63x32; FormatPattern s99.99
      ProcessValue <- "ModbusBuffer_BufferINOut_LookupTable_PinB"
   TextField "Text field_3" at 78,192 size 45x20; Text 'Pfwd:'
   IOField "I/O field_3" at 122,186 size 59x32; FormatPattern 99.99
      ProcessValue <- "ModbusBuffer_BufferINOut_LookupTable_PfwdA"
   IOField "I/O field_4" at 185,186 size 63x32; FormatPattern s99.99
      ProcessValue <- "ModbusBuffer_BufferINOut_LookupTable_PfwdB"
   TextField "Text field_4" at 78,228 size 45x20; Text 'Prev:'
   IOField "I/O field_5" at 122,222 size 59x32; FormatPattern 99.99
      ProcessValue <- "ModbusBuffer_BufferINOut_LookupTable_PrevA"
   IOField "I/O field_6" at 185,222 size 63x32; FormatPattern s99.99
      ProcessValue <- "ModbusBuffer_BufferINOut_LookupTable_PrevB"
   TextField "Text field_9" at 340,224 size 16x25; Text 'P'
   TextField "Text field_12" at 351,234 size 21x14; Text 'REV'
   IOField "Template_I/O Pin dBm" at 372,228 size 50x20; FormatPattern 999.9
      Visibility <- "ModbusBuffer_BufferINOut_SetupData_dBm_unit"
      ProcessValue <- "ModbusBuffer_BufferINOut_CalculatedData_Prev_dBm"
   SymbolicIOField "Template_Symbolic I/O Underrange" at 372,228 size 22x20; TextOn '1'; TextOff '0'; TextList "Text_list_underrange"
      ProcessValue <- "PrevUR"

screen "System information" 480x272, template "Template"
   on GenerateScreen: SetTag("Tag_ScreenNumber", 5)
   TextField "HmiScreenItemData" at 68,78 size 158x20; Text 'HMI device type:'
   TextField "HmiScreenItemData_1" at 230,78 size 246x20; Text 'KTP400 Basic+ PN 15.1.0.0'
   TextField "HmiScreenItemData_2" at 68,99 size 158x20; Text 'Connection:'
   TextField "HmiScreenItemData_3" at 230,99 size 246x20; Text 'PROFINET (X1)'
   TextField "HmiScreenItemData_4" at 68,120 size 158x20; Text 'PLC:'
   TextField "HmiScreenItemData_5" at 230,120 size 246x20; Text 'SIMATIC S7 1200'
   Button "Back" at 65,46 size 136x30; TextOff 'Back'
      on Release: ActivateScreen("System screens", 0)
   TextField "HmiScreenItemData_6" at 69,143 size 158x20; Text 'Program Version:'
   TextField "HmiScreenItemData_7" at 231,143 size 246x20; Text '1.0.0 2025-01-30'

Template "Template_noPrev" 480x272
   TextField "Template_Text field_1" at 94,6 size 23x37; Text 'P'
   TextField "Template_Text field_3" at 109,23 size 30x17; Text 'FWD'
   Button "Alarms" at 1,46 size 63x44; TextOn 'Alarms'; TextOff 'Alarms'; PictureOn "AlarmDisplay_KTP400_Basic_PN_TR"; PictureOff "AlarmDisplay_KTP400_Basic_PN_TR"
      on Release: function_ef3f5d25("Alarm window_Unacknowledged", -1)
   Button "Start screen" at 1,226 size 63x44; TextOn 'Start screen'; TextOff 'Start screen'; PictureOn "NavigateHome_KTP400_Basic_PN_TR"; PictureOff "NavigateHome_KTP400_Basic_PN_TR"
      on Release: ActivateScreen("Root screen", 0)
   GraphicView "Logo" at 0,0 size 94x45; Picture "Logo of HMI_1"
   Button "Template_Button_3" at 1,91 size 63x44; TextOff 'System'
      on Release: ActivateScreen("System screens", 0)
   Group "Group" at 94,6 size 45x37
   IOField "Template_I/O Pfwd" at 142,6 size 80x39; FormatPattern 999
      Visibility <- "ModbusBuffer_BufferINOut_SetupData_dBm_unit"
      ProcessValue <- "AnalogInputs_Pfwd_AnalogIN_Out"
   Switch "Template_Switch_1" at 1,136 size 64x44; TextOn 'Rem'; CaptionText 'Switch'; TextOff 'Loc'
      ProcessValue <- "ModbusBuffer_BufferINOut_SetupData_RemoteMode"
   Switch "Template_Switch_2" at 1,181 size 63x44; TextOn 'dBm'; CaptionText 'Switch'; TextOff 'W'
      ProcessValue <- "ModbusBuffer_BufferINOut_SetupData_dBm_unit"
   SymbolicIOField "Template_Symbolic I/O field_1" at 225,15 size 50x28; TextOn '1'; TextOff '0'; TextList "Text_list_EGU"
      ProcessValue <- "ModbusBuffer_BufferINOut_SetupData_dBm_unit"
   IOField "Template_I/O Pfwd dBm" at 142,6 size 80x39; FormatPattern 999.9
      ProcessValue <- "ModbusBuffer_BufferINOut_CalculatedData_Pfwd_dBm"
      Visibility <- "ModbusBuffer_BufferINOut_SetupData_dBm_unit"
   SymbolicIOField "Symbolic I/O Underrange Pfwd" at 140,5 size 22x39; TextOn '1'; TextOff '0'; TextList "Text_list_underrange"
      ProcessValue <- "PfwdUR"
*)